(* Logix 5000 project; controller PLC_MCC1300_75F1 vendor 1 type 14 code 166 rev 32.11; software revision 32.04; part 71 of 83 *)
(* tags used below, declared in another part *)
   AUX_tConvoy_SL_NULL : UDT_Convoy_SL;
   AUX_xInitialize : BOOL;
   CONST_rgdDestMask : DINT[32];   // Destination Mask
   CONST_tPlant : UDT_PLANT_CONSTANTS;
   GP_TrackingGetFirstPlateInConveyor : GP_TrackingGetFirstPlateInConveyor;
   GP_TrackingPresencePlate : GP_TrackingPresencePlate;
   GP_TrackingSearchPlate : GP_TrackingSearchPlate;
   M310Popup : MAC_Popup_ZC[2];
   M350_M1_DR : AXIS_CIP_DRIVE;
   M350_xReqStopPrevConvForPos : BOOL;
   M350Popup : MAC_Popup_ZC;
   M350Popup_HMW : MAC_Popup_ZC_HMW;
   M350Popup_ReentryCap : UDT_ConvoyCap_ZC;
   M350Popup_SL_DATA : UDT_Convoy_SL;
   M350Popup_xDrivePosEnable : BOOL;
   M350Popup_xQualityComing : BOOL;
   TMP_d : DINT;
   TMP_dBaryc_ins_max : DINT;
   TMP_dBaryc_ins_min : DINT;
   TMP_dIndex : DINT;
   TMP_dIndex2 : DINT;
   TMP_dIndex3 : DINT;
   TMP_dMaskAllowed : DINT;
   TMP_dStartSearch : DINT;
   TMP_dStopSearch : DINT;
   TMP_StartPlusLength : DINT;
   TMP_xAllCullet : BOOL;
   TMP_xAllLiteToCullet : BOOL;
   TMP_xAtLeastOneForQuality : BOOL;
   TMP_xAtLeastOneForSideLeg : BOOL;
   TMP_xDummy : BOOL;
   TMP_xPosHead : BOOL;
   xAlwaysOFF : BOOL;
   xDebugOFF : BOOL;
   Z300_BufferPlate : UDT_LINE_BUFFER_PLATE;
   Z300_Conveyor : UDT_StandConv[29];
   Z300_Conveyor_ALM : MAC_Conveyor_ZC_ALM[29];
   Z300_Conveyor_IN_MOTION : MAC_Conveyor_ZC_IN_MOTION[29];
   Z300_Conveyor_OUT_MOTION : MAC_Conveyor_ZC_OUT_MOTION[29];
   Z300_LineTracking : UDT_LINE_TRACKING;
   Z301 : MAC_Zone_ML;
(* MainProgram, continued *)

   // #####_PRESENCE_PLATE_ON_POPUP_AFTER_POSITIONING_#####
   47: NOP();
   // Search on whole popup size
   48: ADD(150000,M350Popup.AUX_dEndPosition_cmm,TMP_d)GP_TrackingSearchPlate(GP_TrackingSearchPlate,TMP_d,M350Popup.AUX_dStartPosition_cmm,0,Z300_LineTracking,M350Popup.tSearchPlateStop,CONST_tPlant.dNumOfConveyors,CONST_tPlant.dNumCapsConveyor,Z300_BufferPlate);
   49: XIC(M350Popup.tSearchPlateStop.xHeadPresence)MOV(M350Popup.tSearchPlateStop.rgdHeadPointer[0],M350Popup.AUX_dIndexPlateStop);
   50: XIO(M350Popup.tSearchPlateStop.xHeadPresence)XIC(M350Popup.tSearchPlateStop.xTailPresence)MOV(M350Popup.tSearchPlateStop.rgdTailPointer[0],M350Popup.AUX_dIndexPlateStop);
   51: [XIO(M350Popup.tSearchPlateStop.xHeadPresence) XIO(M350Popup.tSearchPlateStop.xTailPresence) ,XIC(Z300_Conveyor[21].ST_xCleaningEnabled) ]MOV(0,M350Popup.AUX_dIndexPlateStop);
   52: [XIC(M350Popup.tSearchPlateStop.xHeadPresence) ,XIC(M350Popup.tSearchPlateStop.xTailPresence) ][OTU(TMP_xAtLeastOneForSideLeg) ,OTU(TMP_xAtLeastOneForQuality) ,OTL(TMP_xAllLiteToCullet) ];
   53: [XIC(M350Popup.tSearchPlateStop.xHeadPresence) ,XIC(M350Popup.tSearchPlateStop.xTailPresence) ]JSR(sbrCheckConvoyZCDestination,5,M350Popup.AUX_dIndexPlateStop,M350Popup.AUX_dDestMaskOppOpSide,CONST_rgdDestMask[24],TMP_xAtLeastOneForQuality,TMP_xAllLiteToCullet,TMP_xAtLeastOneForQuality,TMP_xAllLiteToCullet)XIC(TMP_xAtLeastOneForQuality)[EQU(M350Popup.AUX_dIndexPositioning,M350Popup.AUX_dIndexPlateStop) ,EQU(M350Popup.AUX_dIndexPlatePositioned,M350Popup.AUX_dIndexPlateStop) ,XIO(xDebugOFF) ]OTE(M350Popup.ST_xPlateStopToPopup);
   54: XIO(xAlwaysOFF)XIC(Z300_Conveyor[21].OUTPUT_xPositioning.0)OTE(Z300_Conveyor[21].xReqBypassEndStop);
   55: [XIC(M350Popup.AUX_tSearchPlateData.xPlateHooked) [XIC(M350Popup.tSearchPlateStop.xHeadPresence) ,XIC(M350Popup.tSearchPlateStop.xTailPresence) ,EQU(M350Popup.AUX_dIndexPositioning,Z300_LineTracking.rgtTrkConv[21].Cap[0].dPointer) ] [XIC(TMP_xPosHead) MOV(M350Popup.AUX_dIndexPositioning,TMP_dIndex) [XIC(Z300_BufferPlate.rgtPlate[TMP_dIndex].tData.tFlag.tConveyor.xDoneHeadPositioning) ,XIO(xDebugOFF) XIC(Z300_Conveyor[21].OUTPUT_xPositioning.0) XIC(Z300_Conveyor_OUT_MOTION[21].DR_MAM_M[0].PC) ] ,XIO(TMP_xPosHead) MOV(M350Popup.AUX_dIndexPositioning,TMP_dIndex) XIC(Z300_BufferPlate.rgtPlate[TMP_dIndex].tData.tFlag.tConveyor.xDoneTailPositioning) ] XIC(M350Popup.ST_xPlateStopToPopup) ,XIO(M350Popup.INPUT_xPopupLow) ,XIC(M310Popup[0].ST_xStopPreviousConveyor) ]OTE(Z300_Conveyor[21].xReqStop);
   // Stop tracking update while ending positioning
   56: XIO(xDebugOFF)XIC(M350Popup.AUX_tSearchPlateData.xPlateHooked)MOV(M350Popup.AUX_dIndexPositioning,TMP_dIndex)XIC(M350Popup_xDrivePosEnable)XIO(M350_M1_DR.Registration1InputStatus)ADD(Z300_LineTracking.rgtTrkConv[21].dStartPosition_cmm,Z300_Conveyor[21].AUX_rgdTarget_cmm[0],TMP_d)SUB(TMP_d,Z300_LineTracking.rgtTrkConv[21].dActualRamp_cmm[0],TMP_d)GEQ(Z300_BufferPlate.rgtPlate[TMP_dIndex].tTracking.dPositionHead_cmm,TMP_d)XIC(M350Popup.ST_xPlateStopToPopup)XIC(Z300_Conveyor_IN_MOTION[21].DR_MAM_M[0].IP)XIO(Z300_Conveyor_IN_MOTION[21].DR_MAM_M[0].PC)XIO(Z300_Conveyor_IN_MOTION[21].DR_MAM_M[0].ER)[OTE(Z300_BufferPlate.rgtPlate[TMP_dIndex].tTracking.xHoldAdvancement) ,ADD(M350Popup.AUX_dPosPhotocell_cmm,Z300_Conveyor[21].AUX_rgdTarget_cmm[0],TMP_d) JSR(sbrUpdateTrackingConvoyPosition,2,TMP_dIndex,TMP_d) ];
   57: XIO(xDebugOFF)XIC(Z300_BufferPlate.rgtPlate[TMP_dIndex].tTracking.xHoldAdvancement)GRT(Z300_BufferPlate.rgtPlate[TMP_dIndex].tTracking.dNextCapIndex,0)MOV(Z300_BufferPlate.rgtPlate[TMP_dIndex].tTracking.dNextCapIndex,TMP_dIndex2)OTE(Z300_BufferPlate.rgtPlate[TMP_dIndex2].tTracking.xHoldAdvancement);
   58: XIO(xDebugOFF)XIC(Z300_BufferPlate.rgtPlate[TMP_dIndex2].tTracking.xHoldAdvancement)GRT(Z300_BufferPlate.rgtPlate[TMP_dIndex2].tTracking.dNextCapIndex,0)MOV(Z300_BufferPlate.rgtPlate[TMP_dIndex2].tTracking.dNextCapIndex,TMP_dIndex3)OTE(Z300_BufferPlate.rgtPlate[TMP_dIndex3].tTracking.xHoldAdvancement);
   // Stop previous conveyoy when plate tail has left previous conveyor
   59: XIC(M350Popup.AUX_tSearchPlateData.xPlateHooked)XIC(Z300_LineTracking.rgtTrkConv[21].xGlassPresence)MOV(M350Popup.AUX_dIndexPositioning,TMP_dIndex)[LES(Z300_BufferPlate.rgtPlate[TMP_dIndex].tData.dTotalCaps,2) ,XIO(xDebugOFF) ]XIC(M350Popup_xDrivePosEnable)XIO(M350_M1_DR.Registration1InputStatus)[ADD(Z300_LineTracking.rgtTrkConv[21].dStartPosition_cmm,Z300_Conveyor[21].AUX_rgdTarget_cmm[0],TMP_d) SUB(TMP_d,Z300_LineTracking.rgtTrkConv[21].dActualRamp_cmm[0],TMP_d) GEQ(Z300_BufferPlate.rgtPlate[TMP_dIndex].tTracking.dPositionHead_cmm,TMP_d) ,ADD(Z300_LineTracking.rgtTrkConv[21].dStartPosition_cmm,Z300_BufferPlate.rgtPlate[TMP_dIndex].tData.rgtCap[0].dConvTotLength_cmm,TMP_StartPlusLength) GEQ(Z300_BufferPlate.rgtPlate[TMP_dIndex].tTracking.dPositionHead_cmm,TMP_StartPlusLength) ]OTE(M350_xReqStopPrevConvForPos);
   // #####_PRESENCE_PLATE_UNDER_POPUP_#####
   60: NOP();
   61: ADD(M350Popup.AUX_dStartPosition_cmm,20000,TMP_d)GP_TrackingPresencePlate(GP_TrackingPresencePlate,TMP_d,M350Popup.AUX_dEndPosition_cmm,0,Z300_LineTracking,M350Popup.ST_xPlateUnderPopup);
   62: XIC(M350Popup.AUX_tSearchPlateData.xPlateHooked)GRT(M350Popup.AUX_dIndexPositioning,0)MOV(M350Popup.AUX_dIndexPositioning,TMP_dIndex)[XIC(TMP_xPosHead) GEQ(Z300_BufferPlate.rgtPlate[TMP_dIndex].tTracking.dPositionHead_cmm,M350Popup.AUX_tSearchPlateData.dPositionStopHooked_cmm) ,XIO(TMP_xPosHead) GEQ(Z300_BufferPlate.rgtPlate[TMP_dIndex].tTracking.dPositionTail_cmm,M350Popup.AUX_tSearchPlateData.dPositionStopHooked_cmm) ][OSR(M350Popup.AUX_tSearchPlateData.OSR_xPlateOutHooked,M350Popup.AUX_tSearchPlateData.OS_xPlateOutHooked) ,OTE(M350Popup.ST_xPopupChangeDest) ];
   // Allowed mask calculation for redestination
   63: CPT(TMP_dMaskAllowed,CONST_rgdDestMask[2] OR CONST_rgdDestMask[3]);
   // #####_Change_Destination_#####
   64: XIC(M350Popup.ST_xPopupChangeDest)[JSR(sbrRedestConvoyCapZC,5,M350Popup.AUX_dIndexPositioning,M350Popup.AUX_dDestMaskOpSide,TMP_dMaskAllowed,0,CONST_rgdDestMask[24]) ,OTU(M350Popup.AUX_tSearchPlateData.xPlateHooked) ,OTU(M350Popup_xQualityComing) ,MOV(0,M350Popup.AUX_dIndexPositioning) ,MOV(0,M350Popup.AUX_dIndexPlatePositioned) ];
   65: [XIC(M350Popup.AUX_tSearchPlateData.OS_xPlateOutHooked) ,XIC(M350Popup.AUX_tSearchPlateData.xPlateHooked) XIO(M350Popup.AUX_tSearchPlateData.xIndexCons) ,XIC(Z300_Conveyor[21].ST_xCleaningEnabled) ][MOV(0,M350Popup.AUX_dIndexPositioning) ,OTU(M350Popup.AUX_tSearchPlateData.xPlateHooked) ,OTU(M350Popup_xQualityComing) ];
   // Check if there is a cap destined to popup during a restart of the CPU and make redestination
   66: [XIC(AUX_xInitialize) ,XIC(M350Popup.ST_xPlateInPositionToRise) XIC(M350_M1_DR.Registration1InputStatus) ]XIC(M350Popup.ST_xPlateStopToPopup)GP_TrackingGetFirstPlateInConveyor(GP_TrackingGetFirstPlateInConveyor,Z300_LineTracking.rgtTrkConv[21],CONST_tPlant.dNumCapsConveyor,GP_TrackingGetFirstPlateInConveyor.OUT_dIndex,GP_TrackingGetFirstPlateInConveyor.OUT_dHeadPos)GRT(GP_TrackingGetFirstPlateInConveyor.OUT_dIndex,0)GRT(GP_TrackingGetFirstPlateInConveyor.OUT_dHeadPos,M350Popup.AUX_dStartPosition_cmm)LES(GP_TrackingGetFirstPlateInConveyor.OUT_dHeadPos,M350Popup.AUX_dEndPosition_cmm)MOV(GP_TrackingGetFirstPlateInConveyor.OUT_dIndex,M350Popup.AUX_dIndexPlatePositioned)OTE(M350Popup.OS_xChangeDestAfterRestart);
   // Change destination aftet restart
   67: XIC(M350Popup.OS_xChangeDestAfterRestart)[JSR(sbrRedestConvoyCapZC,5,M350Popup.AUX_dIndexPlatePositioned,M350Popup.AUX_dDestMaskOpSide,TMP_dMaskAllowed,0,CONST_rgdDestMask[24]) ,JSR(sbrTrackingIndexTailConvoy,1,M350Popup.AUX_dIndexPlatePositioned,M350Popup.AUX_dIndexPlateFree) ,OTU(M350Popup.AUX_tSearchPlateData.xPlateHooked) ,OTU(M350Popup_xQualityComing) ,MOV(0,M350Popup.AUX_dIndexPositioning) ,MOV(0,M350Popup.AUX_dIndexPlatePositioned) ];
   68: NOP();
   // #####_Lifting_#####
   69: NOP();
   // Plate in position to raise
   70: XIO(Z300_Conveyor[21].ST_xCleaningEnabled)[XIC(M350Popup.AUX_tSearchPlateData.xPlateHooked) GRT(M350Popup.AUX_dIndexPositioning,0) MOV(M350Popup.AUX_dIndexPositioning,TMP_dIndex) [XIC(TMP_xPosHead) [XIC(Z300_BufferPlate.rgtPlate[TMP_dIndex].tData.tFlag.tConveyor.xDoneHeadPositioning) ,XIC(Z300_Conveyor[21].OUTPUT_xPositioning.0) XIC(Z300_Conveyor_OUT_MOTION[21].DR_MAM_M[0].PC) ] ,XIO(TMP_xPosHead) XIC(Z300_BufferPlate.rgtPlate[TMP_dIndex].tData.tFlag.tConveyor.xDoneTailPositioning) ] XIC(Z300_Conveyor[21].xReqStop) ,XIC(M350Popup.ST_xPlateInPositionToRise) ]XIC(M350Popup.ST_xPlateStopToPopup)XIO(Z300_Conveyor[21].INPUT_xDriveDeceleration.0)XIO(Z300_Conveyor[21].INPUT_xDriveFeedback.0)XIO(M350Popup.ST_xRequestRise)[OTE(M350Popup.ST_xPlateInPositionToRise) ,EQU(M350Popup.AUX_dIndexPlatePositioned,0) MOV(M350Popup.AUX_dIndexPositioning,M350Popup.AUX_dIndexPlatePositioned) ];
   // Request rise
   71: XIO(Z300_Conveyor[21].OUTPUT_xPositioning.0)XIO(M350_M1_DR.Registration1InputStatus)XIC(M350Popup.AUX_tSearchPlateData.xPlateHooked)XIC(M350Popup.ST_xPlateInPositionToRise)[XIC(M350Popup.ST_xPlateToSinglePositioning) ,XIC(M350Popup.ST_xConvoyPositioning) ]XIC(M350Popup.ST_xInitialConditionForRise)XIO(M350Popup.INPUT_xPopupHigh)OTE(M350Popup.ST_xRequestRise);
   // #####_Plate_ready_to_descend_#####
   72: JSR(sbrCheckConvoySLDestination,3,M350Popup_SL_DATA,CONST_rgdDestMask[29],CONST_rgdDestMask[24],TMP_xAllCullet,TMP_xAtLeastOneForQuality);
   // #####_Descending_#####
   73: XIO(Z300_Conveyor[21].OUTPUT_xPositioning.0)XIO(Z300_Conveyor[21].ST_xCleaningEnabled)LEQ(Z301.AUX_dBarPositionCleaning,2620000)XIC(M350Popup.ST_xInitialConditionForDescend)XIO(M350Popup.ST_xPhasesInProgress)[XIO(M350Popup.ST_xPlateUnderPopup) ,XIO(xAlwaysOFF) ][EQU(M350Popup_SL_DATA.rgtCap[0].dID,0) XIO(M350Popup.ST_xPlatePresence) XIO(M350Popup.ST_xPlatePresentOnPopup) ,[XIC(M350Popup.ST_xPlatePresence) ,XIC(M350Popup.ST_xPlatePresentOnPopup) ] [XIO(TMP_xAtLeastOneForQuality) ,XIC(TMP_xAllCullet) ] ][XIO(Z300_LineTracking.rgtTrkConv[21].xGlassPresCom) ,XIC(M350Popup.ST_xPlateToSingleComing) ,XIC(M350Popup.ST_xConvoyComing) ,XIO(xAlwaysOFF) XIC(M350Popup.INPUT_xPopupHigh) ]XIO(M350Popup.INPUT_xPopupLow)OTE(M350Popup.ST_xRequestDescend);
   // #####_Move data to Popup_#####
   74: XIC(M350Popup.AUX_tSearchPlateData.xPlateHooked)XIC(M350Popup.PH_xEndRise)[MOV(M350Popup.AUX_dIndexPositioning,TMP_dIndex) MOV(Z300_BufferPlate.rgtPlate[TMP_dIndex].tTracking.dPosition_cmm,M350Popup.AUX_dPosition_cmm) ,JSR(sbrConvDataLineToSL,3,Z300_BufferPlate.rgtPlate[TMP_dIndex].tData,M350Popup_SL_DATA,0,Z300_BufferPlate.rgtPlate[TMP_dIndex].tData,M350Popup_SL_DATA) ,MOV(0,M350Popup.AUX_dPosition_cmm) ,JSR(sbrTrackingDeleteConvoy,1,M350Popup.AUX_dIndexPositioning) ,OTU(M350Popup.AUX_tSearchPlateData.xPlateHooked) ,OTU(M350Popup_xQualityComing) ,MOV(0,M350Popup.AUX_dIndexPositioning) ,MOV(0,M350Popup.AUX_dIndexPlatePositioned) ,OTL(M350Popup.ST_xPlatePresentOnPopup) ,OTU(M350Popup.ST_xPlateToSinglePositioning) ,OTU(M350Popup.ST_xConvoyPositioning) ];
   75: XIC(M350Popup.ST_xPlatePresentOnPopup)OTE(M350Popup.ST_xPlateDataReadyToSend);
   // Convert from Convoy_ZLU to CapConvoy_ZC and Insert in tracking
   76: XIC(M350Popup.PH_xEndDescend)NEQ(M350Popup_SL_DATA.rgtCap[0].dID,0)ADD(Z300_LineTracking.rgtTrkConv[21].dStartPosition_cmm,M350Popup.AUX_dReqTarget_cmm,TMP_d)JSR(sbrResetLinkConvoy,0)MOV(Z300_LineTracking.rgtTrkConv[21].dStartPosition_cmm,TMP_dBaryc_ins_min)MOV(Z300_LineTracking.rgtTrkConv[21].dEndPosition_cmm,TMP_dBaryc_ins_max)JSR(sbrConvDataSLToLine,6,M350Popup_ReentryCap,M350Popup_SL_DATA,0,TMP_d,TMP_dBaryc_ins_min,TMP_dBaryc_ins_max,M350Popup_ReentryCap,M350Popup_SL_DATA)JSR(sbrPutLinkConvoy,0)JSR(sbrTrackingIndexTailConvoy,1,TMP_dIndex,M350Popup.AUX_dIndexPlateFree);
   // Delete plate data
   77: XIC(M350Popup.PH_xEndDescend)COP(AUX_tConvoy_SL_NULL,M350Popup_SL_DATA,1);
   78: XIO(M350Popup.ST_xPlateDataReadyToSend)XIO(M350Popup.INPUT_xPopupHigh)[XIC(M350Popup.ST_xPlatePresence) ,XIC(M350Popup.ST_xPlatePresentOnPopup) ]ONS(M350Popup.OS_xPlateRemovedBySideLeg)[OTU(M350Popup.ST_xPlatePresence) ,COP(AUX_tConvoy_SL_NULL,M350Popup_SL_DATA,1) ,OTU(M350Popup.ST_xPlatePresentOnPopup) ];
   // #####_SATURATION_#####
   79: GRT(M350Popup_HMW.dSaturationSelection,0)XIC(Z301.ST_xCycleON)[[[XIC(Z300_LineTracking.rgtTrkConv[21].xGlassPresence) ,XIC(Z300_LineTracking.rgtTrkConv[21].xGlassPresCom) ] XIO(Z300_Conveyor[21].ST_xRotationFeedback) ,XIO(xAlwaysOFF) XIO(M350Popup.ST_xInitialConditionForRise) ] ,LES(M350Popup_HMW.dSaturationSelection,1) ][[XIC(Z300_LineTracking.rgtTrkConv[20].xGlassPresence) ,XIC(Z300_LineTracking.rgtTrkConv[20].xGlassPresCom) ] XIO(Z300_Conveyor[20].ST_xRotationFeedback) ,LES(M350Popup_HMW.dSaturationSelection,2) ][[XIC(Z300_LineTracking.rgtTrkConv[19].xGlassPresence) ,XIC(Z300_LineTracking.rgtTrkConv[19].xGlassPresCom) ] XIO(Z300_Conveyor[19].ST_xRotationFeedback) ,LES(M350Popup_HMW.dSaturationSelection,3) ]OTE(TMP_xDummy);
   80: XIC(TMP_xDummy)[[XIC(Z300_LineTracking.rgtTrkConv[18].xGlassPresence) ,XIC(Z300_LineTracking.rgtTrkConv[18].xGlassPresCom) ] XIO(Z300_Conveyor[18].ST_xRotationFeedback) ,LES(M350Popup_HMW.dSaturationSelection,4) ][[XIC(Z300_LineTracking.rgtTrkConv[17].xGlassPresence) ,XIC(Z300_LineTracking.rgtTrkConv[17].xGlassPresCom) ] XIO(Z300_Conveyor[17].ST_xRotationFeedback) ,LES(M350Popup_HMW.dSaturationSelection,5) ]OTE(TMP_xDummy);
   81: XIC(TMP_xDummy)XIC(M350Popup.ST_xPlateComingToPopup)[XIC(M350Popup.INPUT_xPopupHigh) ,XIO(Z300_Conveyor[20].ST_xRotationFeedback) XIO(M350Popup.ST_xInitialConditionForRise) XIO(M350Popup.ST_xPlateStopToPopup) XIC(M350Popup.ST_xConditionToStopPrevious) ][XIC(M350Popup.ST_xPlatePresence) XIO(M350Popup.ST_xPlatePresentOnPopup) OTE(M350Popup.ST_xSaturationConditionPrevious) ,XIC(M350Popup.ST_xPlatePresentOnPopup) OTE(M350Popup.ST_xSaturationConditionPopup) ];
   82: XIC(TMP_xDummy)XIC(M350Popup.ST_xPlateComingToPopup)XIC(M350Popup.INPUT_xPopupLow)XIO(M350Popup.ST_xPlatePresence)XIO(M350Popup.ST_xPlatePresentOnPopup)XIC(M350Popup.ST_xPlateStopToPopup)XIC(M350Popup.AUX_tSearchPlateData.xPlateHooked)NEQ(M350Popup.AUX_dIndexPositioning,0)OTE(M350Popup.ST_xSaturationConditionThis);
   83: [XIC(M350Popup.ST_xSaturationConditionPrevious) XIO(M350Popup.ST_xSaturationConditionPopup) XIO(M350Popup.ST_xSaturationConditionThis) ,XIC(M350Popup.ST_xSaturationConditionThis) XIO(M350Popup.ST_xSaturationConditionPrevious) XIO(M350Popup.ST_xSaturationConditionPopup) ,XIC(M350Popup.ST_xSaturationConditionPopup) XIO(M350Popup.ST_xSaturationConditionPrevious) XIO(M350Popup.ST_xSaturationConditionThis) ]XIO(M350Popup.OS_xSaturationOnPrevious)XIO(M350Popup.OS_xSaturationOnThis)XIO(M350Popup.OS_xSaturationOnPopup)XIO(Z300_Conveyor[21].OUTPUT_xPositioning.0)XIO(M350Popup.ST_xRequestRise)[TON(M350Popup.tmON_Saturation,?,?) ,XIC(M350Popup.tmON_Saturation.DN) [XIC(M350Popup.ST_xSaturationConditionPrevious) OTE(M350Popup.OS_xSaturationOnPrevious) ,XIC(M350Popup.ST_xSaturationConditionThis) OTE(M350Popup.OS_xSaturationOnThis) ,XIC(M350Popup.ST_xSaturationConditionPopup) OTE(M350Popup.OS_xSaturationOnPopup) ] ];
   // Allowed mask calculation for redestination
   84: CPT(TMP_dMaskAllowed,CONST_rgdDestMask[0] OR CONST_rgdDestMask[1] OR CONST_rgdDestMask[2] OR CONST_rgdDestMask[3] OR CONST_rgdDestMask[4] OR CONST_rgdDestMask[5] OR CONST_rgdDestMask[6]);
   85: XIC(M350Popup.OS_xSaturationOnPrevious)GRT(M350Popup.AUX_tSearchPlateData.dIndex,0)[JSR(sbrRedestConvoyCapZC,5,M350Popup.AUX_tSearchPlateData.dIndex,M350Popup.AUX_dDestMaskOpSide,TMP_dMaskAllowed,0,CONST_rgdDestMask[24]) ,NEQ(Z300_BufferPlate.rgtPlate[0].tData.rgtCap[0].rgtLite[0].tDestination.rgxMain,CONST_rgdDestMask[29]) JSR(sbrTrackingIndexTailConvoy,1,M350Popup.AUX_tSearchPlateData.dIndex,M350Popup.AUX_dIndexPlateFree) ];
   86: XIC(M350Popup.OS_xSaturationOnThis)XIC(M350Popup.AUX_tSearchPlateData.xPlateHooked)[GRT(M350Popup.AUX_dIndexPlatePositioned,0) ,XIO(xDebugOFF) ][JSR(sbrRedestConvoyCapZC,5,M350Popup.AUX_dIndexPlatePositioned,M350Popup.AUX_dDestMaskOpSide,TMP_dMaskAllowed,0,CONST_rgdDestMask[24]) ,JSR(sbrRedestConvoyCapZC,5,M350Popup.AUX_dIndexPlatePositioned,M350Popup.AUX_dDestMaskOppOpSide,TMP_dMaskAllowed,0,CONST_rgdDestMask[24]) ,JSR(sbrTrackingIndexTailConvoy,1,M350Popup.AUX_dIndexPositioning,M350Popup.AUX_dIndexPlateFree) ,OTU(M350Popup.AUX_tSearchPlateData.xPlateHooked) ,OTU(M350Popup_xQualityComing) ,MOV(0,M350Popup.AUX_dIndexPositioning) ,MOV(0,M350Popup.AUX_dIndexPlatePositioned) ];
   87: XIC(M350Popup.OS_xSaturationOnPopup)JSR(sbrRedestConvoySL,5,M350Popup_SL_DATA,M350Popup.AUX_dDestMaskOpSide,TMP_dMaskAllowed,0,CONST_rgdDestMask[24],M350Popup_SL_DATA);
   // Change destination of plate after popup if still has its destination
   88: ADD(400000,M350Popup.AUX_dEndPosition_cmm,TMP_dStartSearch)ADD(450000,M350Popup.AUX_dEndPosition_cmm,TMP_dStopSearch)GP_TrackingSearchPlate(GP_TrackingSearchPlate,TMP_dStartSearch,TMP_dStopSearch,0,Z300_LineTracking,M350Popup.tSearchPlateChangeDestAfterPopup,CONST_tPlant.dNumOfConveyors,CONST_tPlant.dNumCapsConveyor,Z300_BufferPlate);
   89: XIC(M350Popup.tSearchPlateChangeDestAfterPopup.xHeadPresence)ONS(M350Popup.OSR_xChangeDestAfterPopup)OTE(M350Popup.OS_xChangeDestAfterPopup);
   90: XIC(M350Popup.OS_xChangeDestAfterPopup)MOV(M350Popup.tSearchPlateChangeDestAfterPopup.rgdHeadPointer[0],M350Popup.AUX_dIndexPlateToChangeDestAfterPopup)CPT(TMP_dMaskAllowed,CONST_rgdDestMask[0] OR CONST_rgdDestMask[1] OR CONST_rgdDestMask[2] OR CONST_rgdDestMask[3] OR CONST_rgdDestMask[4] OR CONST_rgdDestMask[5] OR CONST_rgdDestMask[6])JSR(sbrRedestConvoyCapZC,5,M350Popup.tSearchPlateChangeDestAfterPopup.rgdHeadPointer,M350Popup.AUX_dDestMaskOpSide,TMP_dMaskAllowed,0,CONST_rgdDestMask[24]);
   // #####_CLEANING_#####
   91: XIC(Z300_Conveyor[21].ST_xCleaningEnabled)[OTU(M350Popup.PH_xRise) ,OTU(M350Popup.PH_xDescend) ,MOV(0,M350Popup.AUX_dIndexPositioning) ,XIC(M350Popup.INPUT_xPopupLow) [COP(AUX_tConvoy_SL_NULL,M350Popup_SL_DATA,1) ,OTU(M350Popup.ST_xPlatePresence) ,OTU(M350Popup.ST_xPlatePresentOnPopup) ] ];
   92: XIC(M350Popup.INPUT_xPopupHigh)[COP(AUX_tConvoy_SL_NULL,M350Popup_SL_DATA,1) ,OTU(M350Popup.ST_xPlatePresence) ,OTU(M350Popup.ST_xPlatePresentOnPopup) ];
   93: XIC(M350Popup.ST_xMachineAlarm)OTL(Z300_Conveyor_ALM[21].rgxStoppingFault[0].x0);
END_ROUTINE
